// TIA Portal project "SMSS-ENLAB-01-003-1508-012-PLC-B_V13_SP1_1_V17" (V17) (continued)
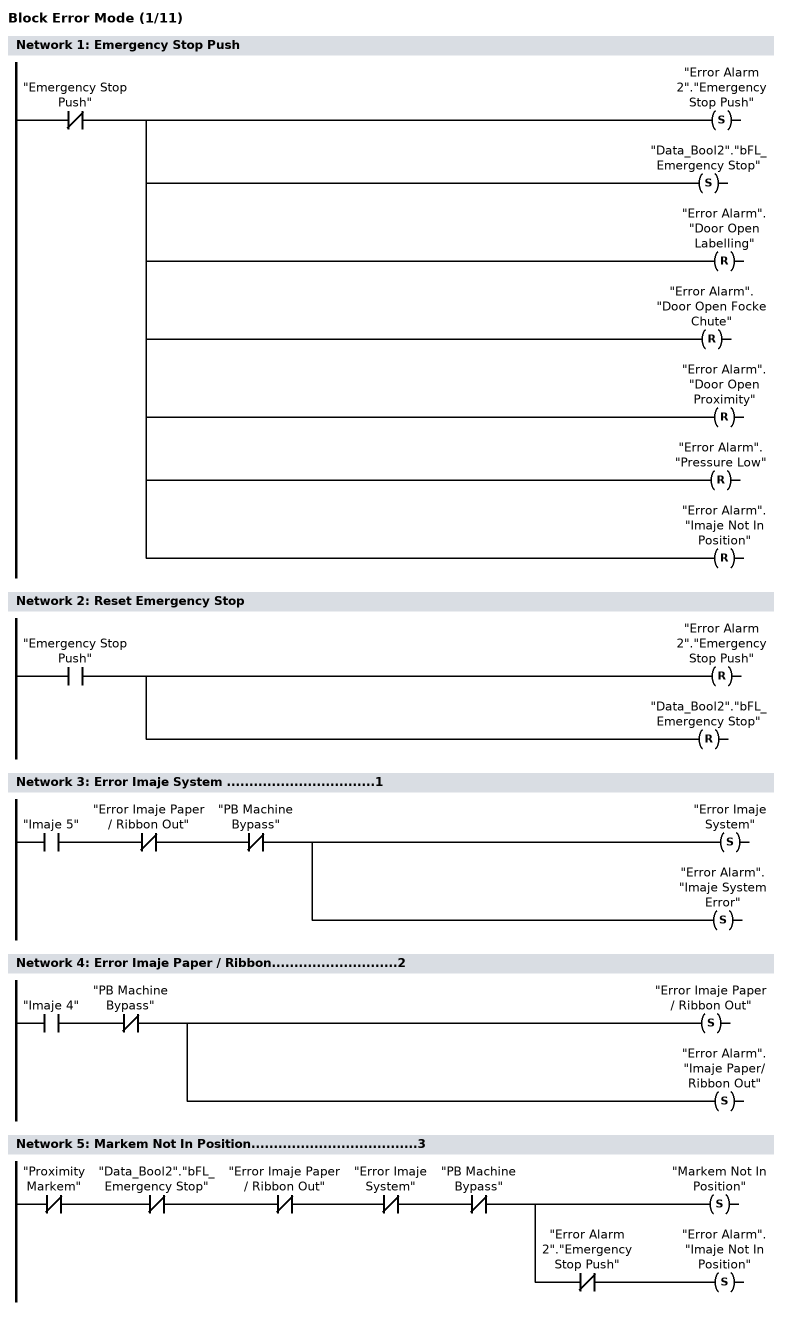
   RUNG wire#powerrail
      I_Contact( "Emergency Stop Push" )
      wire#w1
      S_Coil( "Error Alarm 2"."Emergency Stop Push" )
   END_RUNG
   RUNG wire#w1
      S_Coil( "Data_Bool2"."bFL_Emergency Stop" )
   END_RUNG
   RUNG wire#w1
      R_Coil( "Error Alarm"."Door Open Labelling" )
   END_RUNG
   RUNG wire#w1
      R_Coil( "Error Alarm"."Door Open Focke Chute" )
   END_RUNG
   RUNG wire#w1
      R_Coil( "Error Alarm"."Door Open Proximity" )
   END_RUNG
   RUNG wire#w1
      R_Coil( "Error Alarm"."Pressure Low" )
   END_RUNG
   RUNG wire#w1
      R_Coil( "Error Alarm"."Imaje Not In Position" )
   END_RUNG
   // the same network as SCL:
   IF NOT "Emergency Stop Push" THEN
       "Error Alarm 2"."Emergency Stop Push" := TRUE;
       "Data_Bool2"."bFL_Emergency Stop" := TRUE;
       "Error Alarm"."Door Open Labelling" := FALSE;
       "Error Alarm"."Door Open Focke Chute" := FALSE;
       "Error Alarm"."Door Open Proximity" := FALSE;
       "Error Alarm"."Pressure Low" := FALSE;
       "Error Alarm"."Imaje Not In Position" := FALSE;
   END_IF;
END_REGION

REGION Network 2: Reset Emergency Stop
   RUNG wire#powerrail
      Contact( "Emergency Stop Push" )
      wire#w1
      R_Coil( "Error Alarm 2"."Emergency Stop Push" )
   END_RUNG
   RUNG wire#w1
      R_Coil( "Data_Bool2"."bFL_Emergency Stop" )
   END_RUNG
   // the same network as SCL:
   IF "Emergency Stop Push" THEN
       "Error Alarm 2"."Emergency Stop Push" := FALSE;
       "Data_Bool2"."bFL_Emergency Stop" := FALSE;
   END_IF;
END_REGION

REGION Network 3: Error Imaje System .................................1
   RUNG wire#powerrail
      Contact( "Imaje 5" )
      I_Contact( "Error Imaje Paper / Ribbon Out" )
      I_Contact( "PB Machine Bypass" )
      wire#w1
      S_Coil( "Error Imaje System" )
   END_RUNG
   RUNG wire#w1
      S_Coil( "Error Alarm"."Imaje System Error" )
   END_RUNG
   // the same network as SCL:
   IF "Imaje 5" AND NOT "Error Imaje Paper / Ribbon Out" AND NOT "PB Machine Bypass" THEN
       "Error Imaje System" := TRUE;
       "Error Alarm"."Imaje System Error" := TRUE;
   END_IF;
END_REGION

REGION Network 4: Error Imaje Paper / Ribbon............................2
   RUNG wire#powerrail
      Contact( "Imaje 4" )
      I_Contact( "PB Machine Bypass" )
      wire#w1
      S_Coil( "Error Imaje Paper / Ribbon Out" )
   END_RUNG
   RUNG wire#w1
      S_Coil( "Error Alarm"."Imaje Paper/Ribbon Out" )
   END_RUNG
   // the same network as SCL:
   IF "Imaje 4" AND NOT "PB Machine Bypass" THEN
       "Error Imaje Paper / Ribbon Out" := TRUE;
       "Error Alarm"."Imaje Paper/Ribbon Out" := TRUE;
   END_IF;
END_REGION

REGION Network 5: Markem Not In Position.....................................3
   RUNG wire#powerrail
      I_Contact( "Proximity Markem" )
      I_Contact( "Data_Bool2"."bFL_Emergency Stop" )
      I_Contact( "Error Imaje Paper / Ribbon Out" )
      I_Contact( "Error Imaje System" )
      I_Contact( "PB Machine Bypass" )
      wire#w1
      S_Coil( "Markem Not In Position" )
   END_RUNG
   RUNG wire#w1
      I_Contact( "Error Alarm 2"."Emergency Stop Push" )
      S_Coil( "Error Alarm"."Imaje Not In Position" )
   END_RUNG
   // the same network as SCL:
   #_w1 := NOT "Proximity Markem" AND NOT "Data_Bool2"."bFL_Emergency Stop" AND NOT "Error Imaje Paper / Ribbon Out" AND NOT "Error Imaje System" AND NOT "PB Machine Bypass";
   IF #_w1 THEN "Markem Not In Position" := TRUE; END_IF;
   IF #_w1 AND NOT "Error Alarm 2"."Emergency Stop Push" THEN
       "Error Alarm"."Imaje Not In Position" := TRUE;
   END_IF;
END_REGION

REGION Network 6: Groub Error Imaje Jika baypass mesin Off
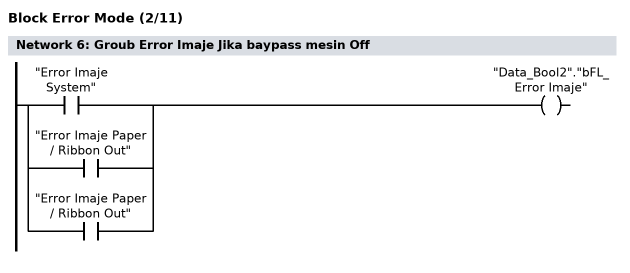
   RUNG wire#powerrail
      Contact( "Error Imaje System" )
      wire#w1
      Coil( "Data_Bool2"."bFL_Error Imaje" )
   END_RUNG
   RUNG wire#powerrail
      Contact( "Error Imaje Paper / Ribbon Out" )
   END_RUNG wire#w1
   RUNG wire#powerrail
      Contact( "Error Imaje Paper / Ribbon Out" )
   END_RUNG wire#w1
   // the same network as SCL:
   "Data_Bool2"."bFL_Error Imaje" := "Error Imaje System" OR "Error Imaje Paper / Ribbon Out" OR "Error Imaje Paper / Ribbon Out";
END_REGION

REGION Network 7: Error Imaje Reset Other Error
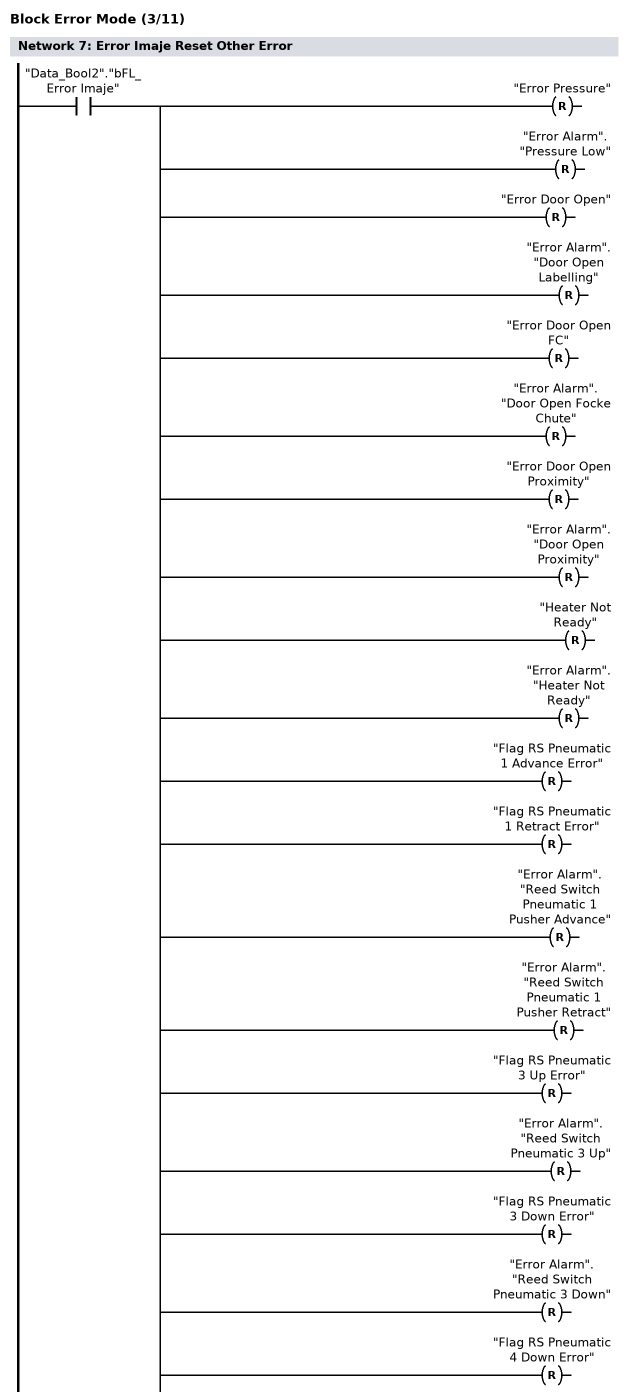
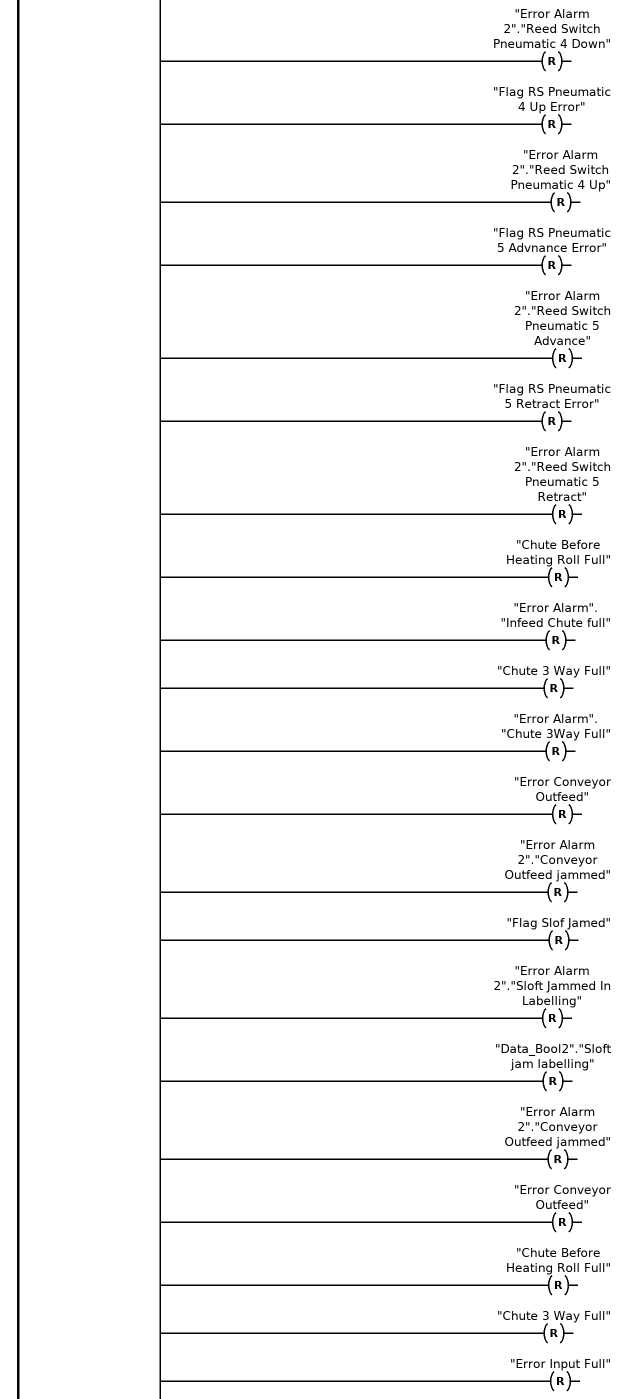
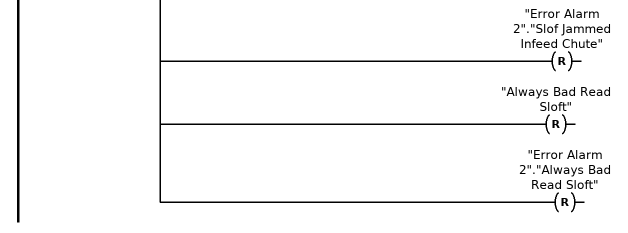
   RUNG wire#powerrail
      Contact( "Data_Bool2"."bFL_Error Imaje" )
      wire#w1
      R_Coil( "Error Pressure" )
   END_RUNG
   RUNG wire#w1
      R_Coil( "Error Alarm"."Pressure Low" )
   END_RUNG
   RUNG wire#w1
      R_Coil( "Error Door Open" )
   END_RUNG
   RUNG wire#w1
      R_Coil( "Error Alarm"."Door Open Labelling" )
   END_RUNG
   RUNG wire#w1
      R_Coil( "Error Door Open FC" )
   END_RUNG
   RUNG wire#w1
      R_Coil( "Error Alarm"."Door Open Focke Chute" )
   END_RUNG
   RUNG wire#w1
      R_Coil( "Error Door Open Proximity" )
   END_RUNG
   RUNG wire#w1
      R_Coil( "Error Alarm"."Door Open Proximity" )
   END_RUNG
   RUNG wire#w1
      R_Coil( "Heater Not Ready" )
   END_RUNG
   RUNG wire#w1
      R_Coil( "Error Alarm"."Heater Not Ready" )
   END_RUNG
   RUNG wire#w1
      R_Coil( "Flag RS Pneumatic 1 Advance Error" )
   END_RUNG
   RUNG wire#w1
      R_Coil( "Flag RS Pneumatic 1 Retract Error" )
   END_RUNG
   RUNG wire#w1
      R_Coil( "Error Alarm"."Reed Switch Pneumatic 1 Pusher Advance" )
   END_RUNG
   RUNG wire#w1
      R_Coil( "Error Alarm"."Reed Switch Pneumatic 1 Pusher Retract" )
   END_RUNG
   RUNG wire#w1
      R_Coil( "Flag RS Pneumatic 3 Up Error" )
   END_RUNG
   RUNG wire#w1
      R_Coil( "Error Alarm"."Reed Switch Pneumatic 3 Up" )
   END_RUNG
   RUNG wire#w1
      R_Coil( "Flag RS Pneumatic 3 Down Error" )
   END_RUNG
   RUNG wire#w1
      R_Coil( "Error Alarm"."Reed Switch Pneumatic 3 Down" )
   END_RUNG
   RUNG wire#w1
      R_Coil( "Flag RS Pneumatic 4 Down Error" )
   END_RUNG
   RUNG wire#w1
      R_Coil( "Error Alarm 2"."Reed Switch Pneumatic 4 Down" )
   END_RUNG
   RUNG wire#w1
      R_Coil( "Flag RS Pneumatic 4 Up Error" )
   END_RUNG
   RUNG wire#w1
      R_Coil( "Error Alarm 2"."Reed Switch Pneumatic 4 Up" )
   END_RUNG
   RUNG wire#w1
      R_Coil( "Flag RS Pneumatic 5 Advnance Error" )
   END_RUNG
   RUNG wire#w1
      R_Coil( "Error Alarm 2"."Reed Switch Pneumatic 5 Advance" )
   END_RUNG
   RUNG wire#w1
      R_Coil( "Flag RS Pneumatic 5 Retract Error" )
   END_RUNG
   RUNG wire#w1
      R_Coil( "Error Alarm 2"."Reed Switch Pneumatic 5 Retract" )
   END_RUNG
   RUNG wire#w1
      R_Coil( "Chute Before Heating Roll Full" )
   END_RUNG
   RUNG wire#w1
      R_Coil( "Error Alarm"."Infeed Chute full" )
   END_RUNG
   RUNG wire#w1
      R_Coil( "Chute 3 Way Full" )
   END_RUNG
   RUNG wire#w1
      R_Coil( "Error Alarm"."Chute 3Way Full" )
   END_RUNG
   RUNG wire#w1
      R_Coil( "Error Conveyor Outfeed" )
   END_RUNG
   RUNG wire#w1
      R_Coil( "Error Alarm 2"."Conveyor Outfeed jammed" )
   END_RUNG
   RUNG wire#w1
      R_Coil( "Flag Slof Jamed" )
   END_RUNG
   RUNG wire#w1
      R_Coil( "Error Alarm 2"."Sloft Jammed In Labelling" )
   END_RUNG
   RUNG wire#w1
      R_Coil( "Data_Bool2"."Sloft jam labelling" )
   END_RUNG
   RUNG wire#w1
      R_Coil( "Error Alarm 2"."Conveyor Outfeed jammed" )
   END_RUNG
   RUNG wire#w1
      R_Coil( "Error Conveyor Outfeed" )
   END_RUNG
   RUNG wire#w1
      R_Coil( "Chute Before Heating Roll Full" )
   END_RUNG
   RUNG wire#w1
      R_Coil( "Chute 3 Way Full" )
   END_RUNG
   RUNG wire#w1
      R_Coil( "Error Input Full" )
   END_RUNG
   RUNG wire#w1
      R_Coil( "Error Alarm 2"."Slof Jammed Infeed Chute" )
   END_RUNG
   RUNG wire#w1
      R_Coil( "Always Bad Read Sloft" )
   END_RUNG
   RUNG wire#w1
      R_Coil( "Error Alarm 2"."Always Bad Read Sloft" )
   END_RUNG
   // the same network as SCL:
   IF "Data_Bool2"."bFL_Error Imaje" THEN
       "Error Pressure" := FALSE;
       "Error Alarm"."Pressure Low" := FALSE;
       "Error Door Open" := FALSE;
       "Error Alarm"."Door Open Labelling" := FALSE;
       "Error Door Open FC" := FALSE;
       "Error Alarm"."Door Open Focke Chute" := FALSE;
       "Error Door Open Proximity" := FALSE;
       "Error Alarm"."Door Open Proximity" := FALSE;
       "Heater Not Ready" := FALSE;
       "Error Alarm"."Heater Not Ready" := FALSE;
       "Flag RS Pneumatic 1 Advance Error" := FALSE;
       "Flag RS Pneumatic 1 Retract Error" := FALSE;
       "Error Alarm"."Reed Switch Pneumatic 1 Pusher Advance" := FALSE;
       "Error Alarm"."Reed Switch Pneumatic 1 Pusher Retract" := FALSE;
       "Flag RS Pneumatic 3 Up Error" := FALSE;
       "Error Alarm"."Reed Switch Pneumatic 3 Up" := FALSE;
       "Flag RS Pneumatic 3 Down Error" := FALSE;
       "Error Alarm"."Reed Switch Pneumatic 3 Down" := FALSE;
       "Flag RS Pneumatic 4 Down Error" := FALSE;
       "Error Alarm 2"."Reed Switch Pneumatic 4 Down" := FALSE;
       "Flag RS Pneumatic 4 Up Error" := FALSE;
       "Error Alarm 2"."Reed Switch Pneumatic 4 Up" := FALSE;
       "Flag RS Pneumatic 5 Advnance Error" := FALSE;
       "Error Alarm 2"."Reed Switch Pneumatic 5 Advance" := FALSE;
       "Flag RS Pneumatic 5 Retract Error" := FALSE;
       "Error Alarm 2"."Reed Switch Pneumatic 5 Retract" := FALSE;
       "Chute Before Heating Roll Full" := FALSE;
       "Error Alarm"."Infeed Chute full" := FALSE;
       "Chute 3 Way Full" := FALSE;
       "Error Alarm"."Chute 3Way Full" := FALSE;
       "Error Conveyor Outfeed" := FALSE;
       "Error Alarm 2"."Conveyor Outfeed jammed" := FALSE;
       "Flag Slof Jamed" := FALSE;
       "Error Alarm 2"."Sloft Jammed In Labelling" := FALSE;
       "Data_Bool2"."Sloft jam labelling" := FALSE;
       "Error Alarm 2"."Conveyor Outfeed jammed" := FALSE;
       "Error Conveyor Outfeed" := FALSE;
       "Chute Before Heating Roll Full" := FALSE;
       "Chute 3 Way Full" := FALSE;
       "Error Input Full" := FALSE;
       "Error Alarm 2"."Slof Jammed Infeed Chute" := FALSE;
       "Always Bad Read Sloft" := FALSE;
       "Error Alarm 2"."Always Bad Read Sloft" := FALSE;
   END_IF;
END_REGION

REGION Network 8: Other Error Imaje Reset Error Imaje
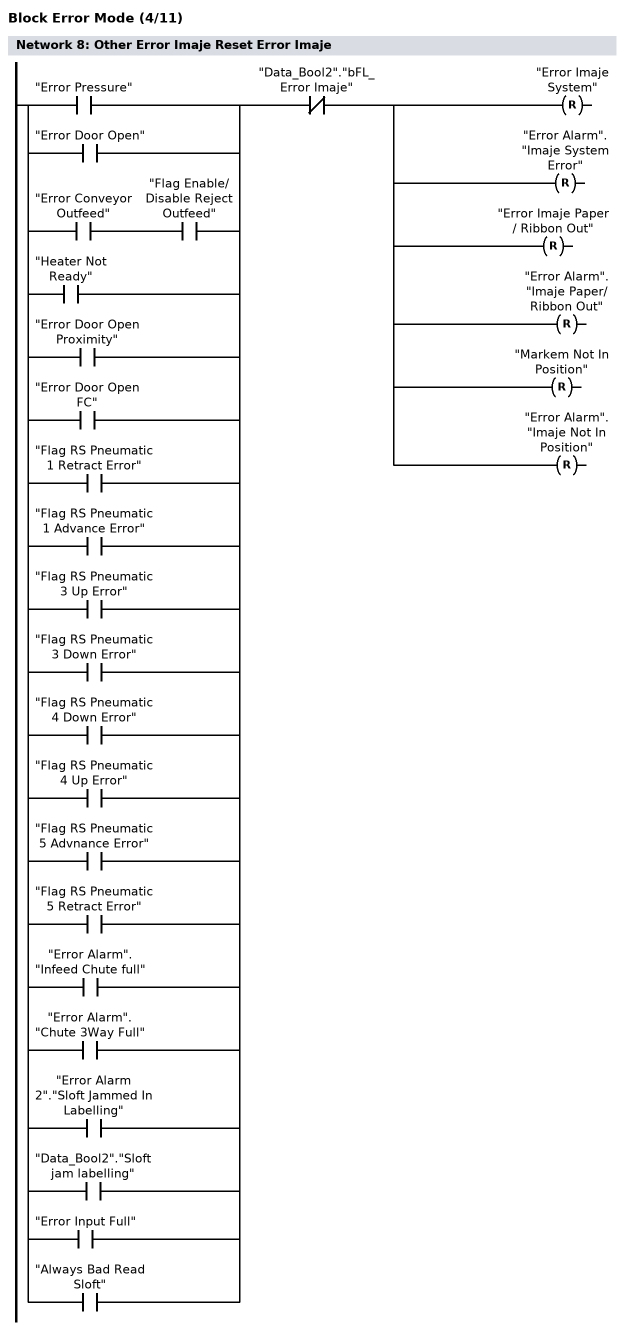
   RUNG wire#powerrail
      Contact( "Error Pressure" )
      wire#w1
      I_Contact( "Data_Bool2"."bFL_Error Imaje" )
      wire#w2
      R_Coil( "Error Imaje System" )
   END_RUNG
   RUNG wire#powerrail
      Contact( "Error Door Open" )
   END_RUNG wire#w1
   RUNG wire#powerrail
      Contact( "Error Conveyor Outfeed" )
      Contact( "Flag Enable/Disable Reject Outfeed" )
   END_RUNG wire#w1
   RUNG wire#powerrail
      Contact( "Heater Not Ready" )
   END_RUNG wire#w1
   RUNG wire#powerrail
      Contact( "Error Door Open Proximity" )
   END_RUNG wire#w1
   RUNG wire#powerrail
      Contact( "Error Door Open FC" )
   END_RUNG wire#w1
   RUNG wire#powerrail
      Contact( "Flag RS Pneumatic 1 Retract Error" )
   END_RUNG wire#w1
   RUNG wire#powerrail
      Contact( "Flag RS Pneumatic 1 Advance Error" )
   END_RUNG wire#w1
   RUNG wire#powerrail
      Contact( "Flag RS Pneumatic 3 Up Error" )
   END_RUNG wire#w1
   RUNG wire#powerrail
      Contact( "Flag RS Pneumatic 3 Down Error" )
   END_RUNG wire#w1
   RUNG wire#powerrail
      Contact( "Flag RS Pneumatic 4 Down Error" )
   END_RUNG wire#w1
   RUNG wire#powerrail
      Contact( "Flag RS Pneumatic 4 Up Error" )
   END_RUNG wire#w1
   RUNG wire#powerrail
      Contact( "Flag RS Pneumatic 5 Advnance Error" )
   END_RUNG wire#w1
   RUNG wire#powerrail
      Contact( "Flag RS Pneumatic 5 Retract Error" )
   END_RUNG wire#w1
   RUNG wire#powerrail
      Contact( "Error Alarm"."Infeed Chute full" )
   END_RUNG wire#w1
   RUNG wire#powerrail
      Contact( "Error Alarm"."Chute 3Way Full" )
   END_RUNG wire#w1
   RUNG wire#powerrail
      Contact( "Error Alarm 2"."Sloft Jammed In Labelling" )
   END_RUNG wire#w1
   RUNG wire#powerrail
      Contact( "Data_Bool2"."Sloft jam labelling" )
   END_RUNG wire#w1
   RUNG wire#powerrail
      Contact( "Error Input Full" )
   END_RUNG wire#w1
   RUNG wire#powerrail
      Contact( "Always Bad Read Sloft" )
   END_RUNG wire#w1
   RUNG wire#w2
      R_Coil( "Error Alarm"."Imaje System Error" )
   END_RUNG
   RUNG wire#w2
      R_Coil( "Error Imaje Paper / Ribbon Out" )
   END_RUNG
   RUNG wire#w2
      R_Coil( "Error Alarm"."Imaje Paper/Ribbon Out" )
   END_RUNG
   RUNG wire#w2
      R_Coil( "Markem Not In Position" )
   END_RUNG
   RUNG wire#w2
      R_Coil( "Error Alarm"."Imaje Not In Position" )
   END_RUNG
   // the same network as SCL:
   IF ("Error Pressure" OR "Error Door Open" OR ("Error Conveyor Outfeed" AND "Flag Enable/Disable Reject Outfeed") OR "Heater Not Ready" OR "Error Door Open Proximity" OR "Error Door Open FC" OR "Flag RS Pneumatic 1 Retract Error" OR "Flag RS Pneumatic 1 Advance Error" OR "Flag RS Pneumatic 3 Up Error" OR "Flag RS Pneumatic 3 Down Error" OR "Flag RS Pneumatic 4 Down Error" OR "Flag RS Pneumatic 4 Up Error" OR "Flag RS Pneumatic 5 Advnance Error" OR "Flag RS Pneumatic 5 Retract Error" OR "Error Alarm"."Infeed Chute full" OR "Error Alarm"."Chute 3Way Full" OR "Error Alarm 2"."Sloft Jammed In Labelling" OR "Data_Bool2"."Sloft jam labelling" OR "Error Input Full" OR "Always Bad Read Sloft") AND NOT "Data_Bool2"."bFL_Error Imaje" THEN
       "Error Imaje System" := FALSE;
       "Error Alarm"."Imaje System Error" := FALSE;
       "Error Imaje Paper / Ribbon Out" := FALSE;
       "Error Alarm"."Imaje Paper/Ribbon Out" := FALSE;
       "Markem Not In Position" := FALSE;
       "Error Alarm"."Imaje Not In Position" := FALSE;
   END_IF;
END_REGION

REGION Network 9: Set Bad Read Berturut-rurut -----------> mesin Error ..................................4
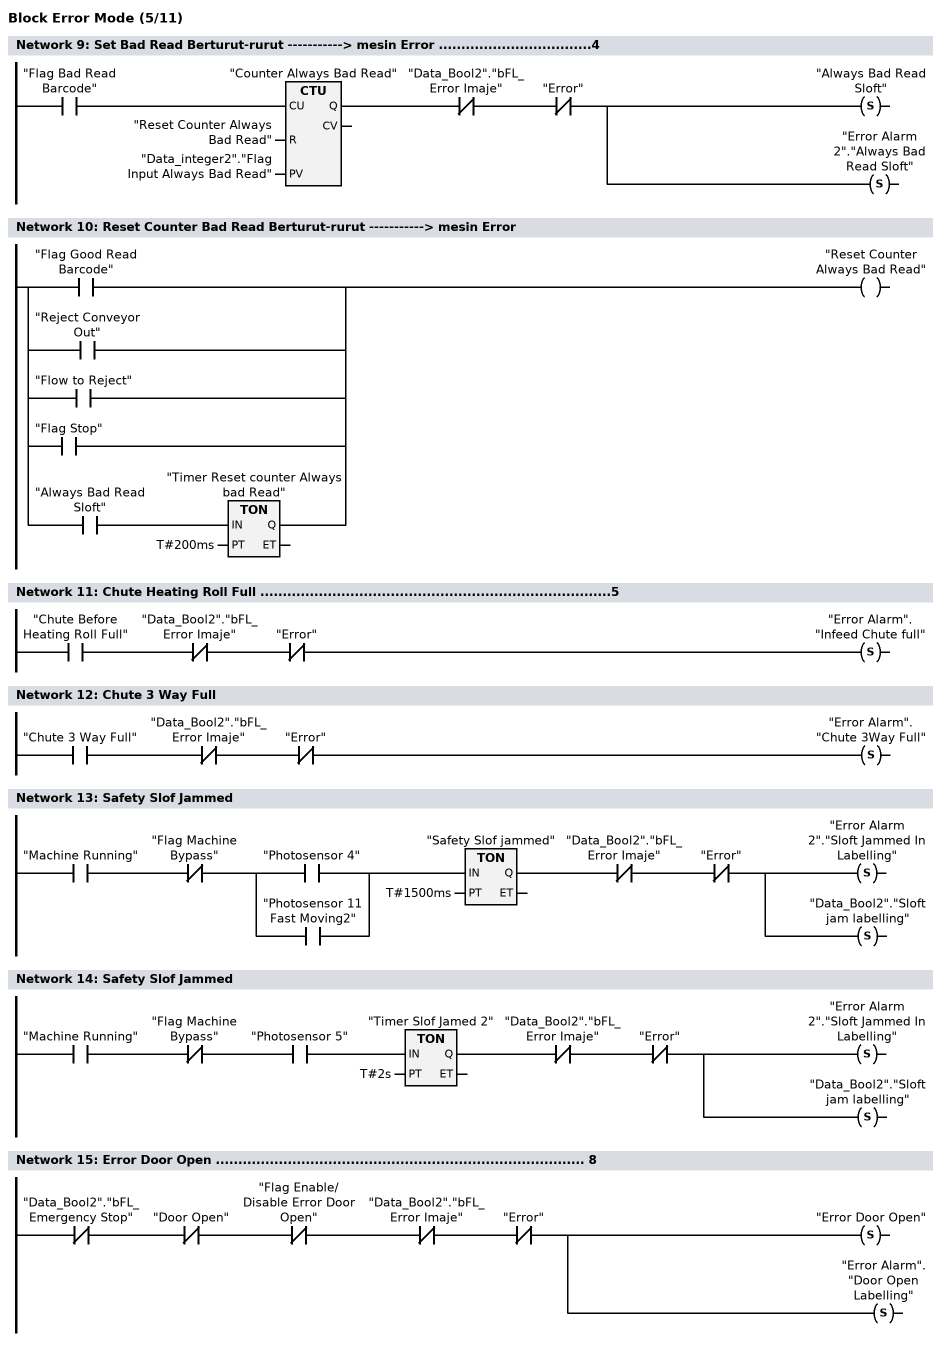
   "Counter Always Bad Read".CTU(CU := "Flag Bad Read Barcode",
                           R := "Reset Counter Always Bad Read",
                           PV := "Data_integer2"."Flag Input Always Bad Read");
   IF "Counter Always Bad Read".Q AND NOT "Data_Bool2"."bFL_Error Imaje" AND NOT "Error" THEN
       "Always Bad Read Sloft" := TRUE;
       "Error Alarm 2"."Always Bad Read Sloft" := TRUE;
   END_IF;
END_REGION

REGION Network 10: Reset Counter Bad Read Berturut-rurut -----------> mesin Error
   "Timer Reset counter Always bad Read".TON(IN := "Always Bad Read Sloft", PT := T#200ms);
   "Reset Counter Always Bad Read" := "Flag Good Read Barcode" OR "Reject Conveyor Out" OR "Flow to Reject" OR "Flag Stop" OR "Timer Reset counter Always bad Read".Q;
END_REGION

REGION Network 11: Chute Heating Roll Full ..............................................................................5
   RUNG wire#powerrail
      Contact( "Chute Before Heating Roll Full" )
      I_Contact( "Data_Bool2"."bFL_Error Imaje" )
      I_Contact( "Error" )
      S_Coil( "Error Alarm"."Infeed Chute full" )
   END_RUNG
   // the same network as SCL:
   IF "Chute Before Heating Roll Full" AND NOT "Data_Bool2"."bFL_Error Imaje" AND NOT "Error" THEN
       "Error Alarm"."Infeed Chute full" := TRUE;
   END_IF;
END_REGION

REGION Network 12: Chute 3 Way Full
   RUNG wire#powerrail
      Contact( "Chute 3 Way Full" )
      I_Contact( "Data_Bool2"."bFL_Error Imaje" )
      I_Contact( "Error" )
      S_Coil( "Error Alarm"."Chute 3Way Full" )
   END_RUNG
   // the same network as SCL:
   IF "Chute 3 Way Full" AND NOT "Data_Bool2"."bFL_Error Imaje" AND NOT "Error" THEN
       "Error Alarm"."Chute 3Way Full" := TRUE;
   END_IF;
END_REGION

REGION Network 13: Safety Slof Jammed
   "Safety Slof jammed".TON(IN := "Machine Running" AND NOT "Flag Machine Bypass" AND ("Photosensor 4" OR "Photosensor 11 Fast Moving2"),
                           PT := T#1500ms);
   IF "Safety Slof jammed".Q AND NOT "Data_Bool2"."bFL_Error Imaje" AND NOT "Error" THEN
       "Error Alarm 2"."Sloft Jammed In Labelling" := TRUE;
       "Data_Bool2"."Sloft jam labelling" := TRUE;
   END_IF;
END_REGION

REGION Network 14: Safety Slof Jammed
   "Timer Slof Jamed 2".TON(IN := "Machine Running" AND NOT "Flag Machine Bypass" AND "Photosensor 5",
                           PT := T#2s);
   IF "Timer Slof Jamed 2".Q AND NOT "Data_Bool2"."bFL_Error Imaje" AND NOT "Error" THEN
       "Error Alarm 2"."Sloft Jammed In Labelling" := TRUE;
       "Data_Bool2"."Sloft jam labelling" := TRUE;
   END_IF;
END_REGION

REGION Network 15: Error Door Open .................................................................................. 8
   RUNG wire#powerrail
      I_Contact( "Data_Bool2"."bFL_Emergency Stop" )
      I_Contact( "Door Open" )
      I_Contact( "Flag Enable/Disable Error Door Open" )
      I_Contact( "Data_Bool2"."bFL_Error Imaje" )
      I_Contact( "Error" )
      wire#w1
      S_Coil( "Error Door Open" )
   END_RUNG
   RUNG wire#w1
      S_Coil( "Error Alarm"."Door Open Labelling" )
   END_RUNG
   // the same network as SCL:
   IF NOT "Data_Bool2"."bFL_Emergency Stop" AND NOT "Door Open" AND NOT "Flag Enable/Disable Error Door Open" AND NOT "Data_Bool2"."bFL_Error Imaje" AND NOT "Error" THEN
       "Error Door Open" := TRUE;
       "Error Alarm"."Door Open Labelling" := TRUE;
   END_IF;
END_REGION

REGION Network 16: Error Door Open FC
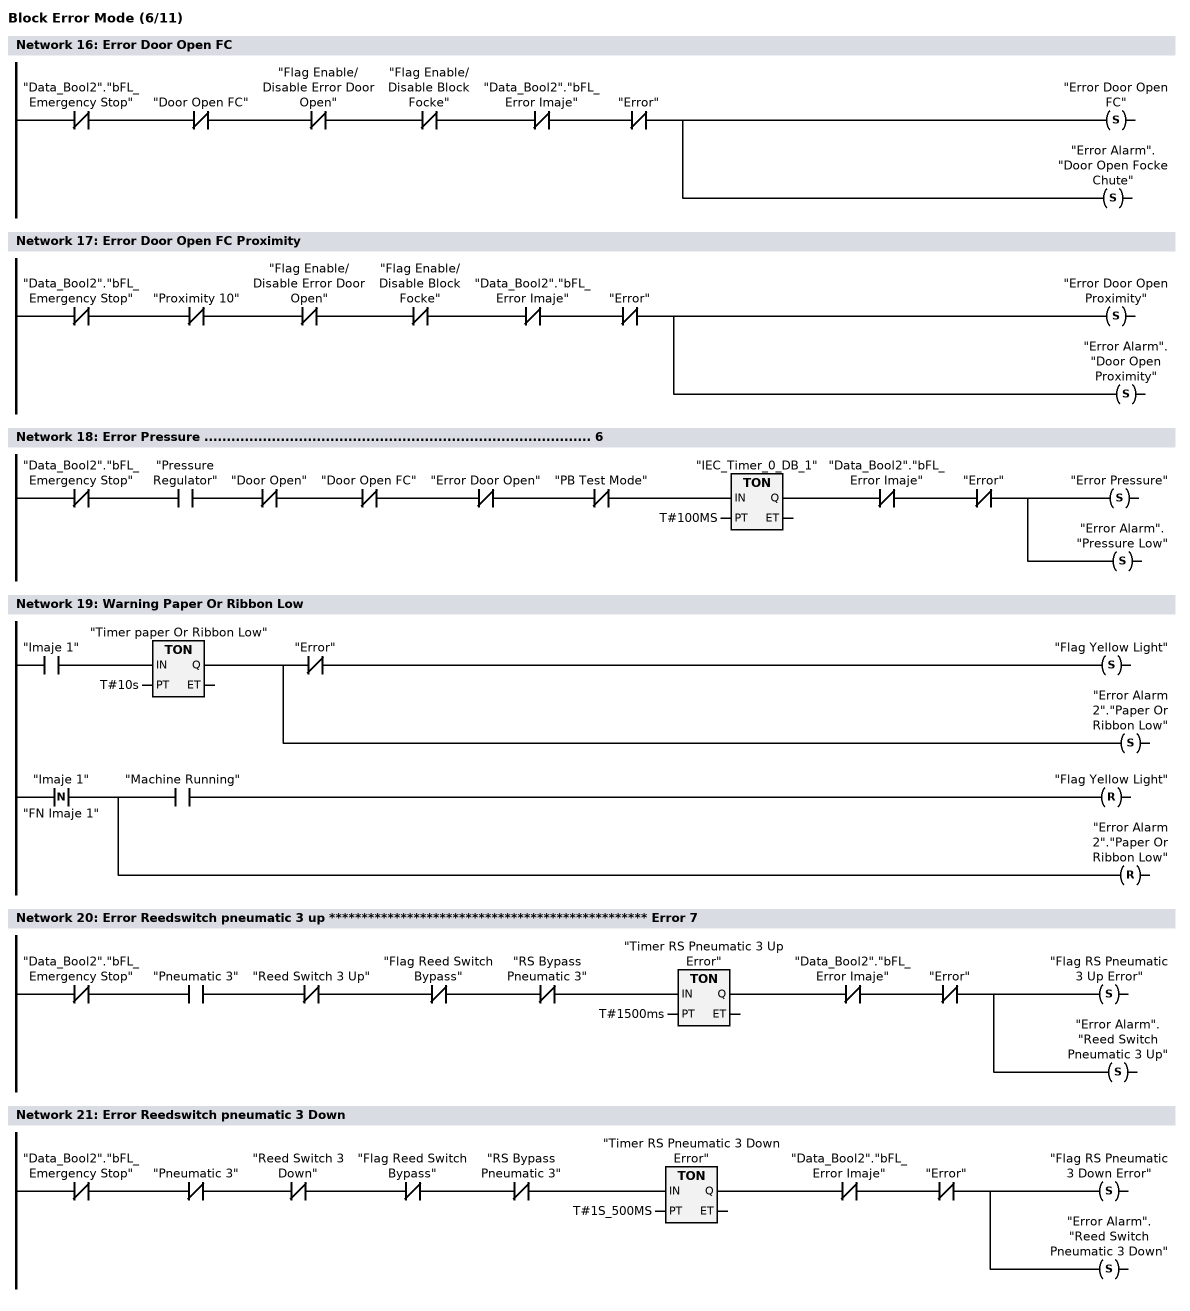
   RUNG wire#powerrail
      I_Contact( "Data_Bool2"."bFL_Emergency Stop" )
      I_Contact( "Door Open FC" )
      I_Contact( "Flag Enable/Disable Error Door Open" )
      I_Contact( "Flag Enable/Disable Block Focke" )
      I_Contact( "Data_Bool2"."bFL_Error Imaje" )
      I_Contact( "Error" )
      wire#w1
      S_Coil( "Error Door Open FC" )
   END_RUNG
   RUNG wire#w1
      S_Coil( "Error Alarm"."Door Open Focke Chute" )
   END_RUNG
   // the same network as SCL:
   IF NOT "Data_Bool2"."bFL_Emergency Stop" AND NOT "Door Open FC" AND NOT "Flag Enable/Disable Error Door Open" AND NOT "Flag Enable/Disable Block Focke" AND NOT "Data_Bool2"."bFL_Error Imaje" AND NOT "Error" THEN
       "Error Door Open FC" := TRUE;
       "Error Alarm"."Door Open Focke Chute" := TRUE;
   END_IF;
END_REGION

REGION Network 17: Error Door Open FC Proximity
   RUNG wire#powerrail
      I_Contact( "Data_Bool2"."bFL_Emergency Stop" )
      I_Contact( "Proximity 10" )
      I_Contact( "Flag Enable/Disable Error Door Open" )
      I_Contact( "Flag Enable/Disable Block Focke" )
      I_Contact( "Data_Bool2"."bFL_Error Imaje" )
      I_Contact( "Error" )
      wire#w1
      S_Coil( "Error Door Open Proximity" )
   END_RUNG
   RUNG wire#w1
      S_Coil( "Error Alarm"."Door Open Proximity" )
   END_RUNG
   // the same network as SCL:
   IF NOT "Data_Bool2"."bFL_Emergency Stop" AND NOT "Proximity 10" AND NOT "Flag Enable/Disable Error Door Open" AND NOT "Flag Enable/Disable Block Focke" AND NOT "Data_Bool2"."bFL_Error Imaje" AND NOT "Error" THEN
       "Error Door Open Proximity" := TRUE;
       "Error Alarm"."Door Open Proximity" := TRUE;
   END_IF;
END_REGION

REGION Network 18: Error Pressure ...................................................................................... 6
   "IEC_Timer_0_DB_1".TON(IN := NOT "Data_Bool2"."bFL_Emergency Stop" AND "Pressure Regulator" AND NOT "Door Open" AND NOT "Door Open FC" AND NOT "Error Door Open" AND NOT "PB Test Mode",
                          PT := T#100MS);
   IF "IEC_Timer_0_DB_1".Q AND NOT "Data_Bool2"."bFL_Error Imaje" AND NOT "Error" THEN
       "Error Pressure" := TRUE;
       "Error Alarm"."Pressure Low" := TRUE;
   END_IF;
END_REGION

REGION Network 19: Warning Paper Or Ribbon Low
   "Timer paper Or Ribbon Low".TON(IN := "Imaje 1", PT := T#10s);
   IF "Timer paper Or Ribbon Low".Q AND NOT "Error" THEN "Flag Yellow Light" := TRUE; END_IF;
   IF "Timer paper Or Ribbon Low".Q THEN "Error Alarm 2"."Paper Or Ribbon Low" := TRUE; END_IF;
   #_w1 := NOT "Imaje 1" AND "FN Imaje 1";   // falling edge of "Imaje 1"
   "FN Imaje 1" := "Imaje 1";
   IF #_w1 AND "Machine Running" THEN "Flag Yellow Light" := FALSE; END_IF;
   IF #_w1 THEN "Error Alarm 2"."Paper Or Ribbon Low" := FALSE; END_IF;
END_REGION

REGION Network 20: Error Reedswitch pneumatic 3 up ************************************************* Error 7
   "Timer RS Pneumatic 3 Up Error".TON(IN := NOT "Data_Bool2"."bFL_Emergency Stop" AND "Pneumatic 3" AND NOT "Reed Switch 3 Up" AND NOT "Flag Reed Switch Bypass" AND NOT "RS Bypass Pneumatic 3",
                           PT := T#1500ms);
   IF "Timer RS Pneumatic 3 Up Error".Q AND NOT "Data_Bool2"."bFL_Error Imaje" AND NOT "Error" THEN
       "Flag RS Pneumatic 3 Up Error" := TRUE;
       "Error Alarm"."Reed Switch Pneumatic 3 Up" := TRUE;
   END_IF;
END_REGION

REGION Network 21: Error Reedswitch pneumatic 3 Down
   "Timer RS Pneumatic 3 Down Error".TON(IN := NOT "Data_Bool2"."bFL_Emergency Stop" AND NOT "Pneumatic 3" AND NOT "Reed Switch 3 Down" AND NOT "Flag Reed Switch Bypass" AND NOT "RS Bypass Pneumatic 3",
                           PT := T#1S_500MS);
   IF "Timer RS Pneumatic 3 Down Error".Q AND NOT "Data_Bool2"."bFL_Error Imaje" AND NOT "Error" THEN
       "Flag RS Pneumatic 3 Down Error" := TRUE;
       "Error Alarm"."Reed Switch Pneumatic 3 Down" := TRUE;
   END_IF;
END_REGION

REGION Network 22: Error Reedswitch pneumatic 4 Down
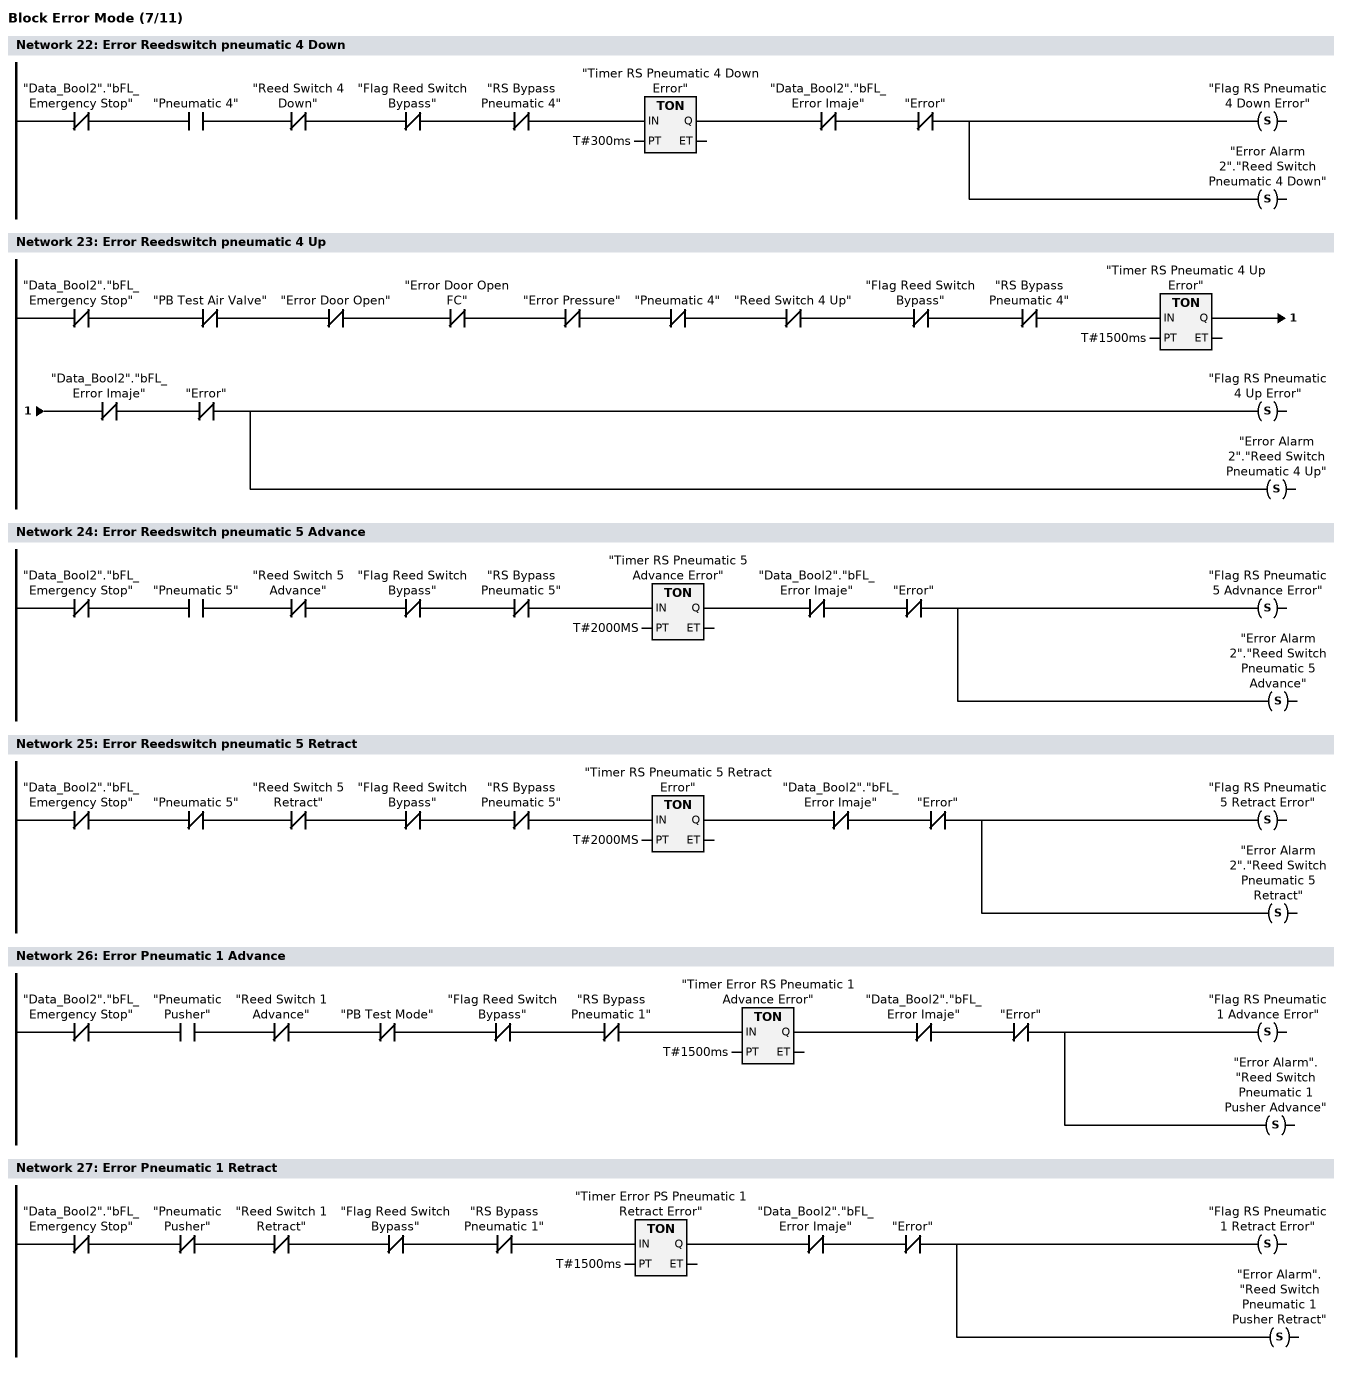
   "Timer RS Pneumatic 4 Down Error".TON(IN := NOT "Data_Bool2"."bFL_Emergency Stop" AND "Pneumatic 4" AND NOT "Reed Switch 4 Down" AND NOT "Flag Reed Switch Bypass" AND NOT "RS Bypass Pneumatic 4",
                           PT := T#300ms);
   IF "Timer RS Pneumatic 4 Down Error".Q AND NOT "Data_Bool2"."bFL_Error Imaje" AND NOT "Error" THEN
       "Flag RS Pneumatic 4 Down Error" := TRUE;
       "Error Alarm 2"."Reed Switch Pneumatic 4 Down" := TRUE;
   END_IF;
END_REGION

REGION Network 23: Error Reedswitch pneumatic 4 Up
   "Timer RS Pneumatic 4 Up Error".TON(IN := NOT "Data_Bool2"."bFL_Emergency Stop" AND NOT "PB Test Air Valve" AND NOT "Error Door Open" AND NOT "Error Door Open FC" AND NOT "Error Pressure" AND NOT "Pneumatic 4" AND NOT "Reed Switch 4 Up" AND NOT "Flag Reed Switch Bypass" AND NOT "RS Bypass Pneumatic 4",
                           PT := T#1500ms);
   IF "Timer RS Pneumatic 4 Up Error".Q AND NOT "Data_Bool2"."bFL_Error Imaje" AND NOT "Error" THEN
       "Flag RS Pneumatic 4 Up Error" := TRUE;
       "Error Alarm 2"."Reed Switch Pneumatic 4 Up" := TRUE;
   END_IF;
END_REGION

REGION Network 24: Error Reedswitch pneumatic 5 Advance
   "Timer RS Pneumatic 5 Advance Error".TON(IN := NOT "Data_Bool2"."bFL_Emergency Stop" AND "Pneumatic 5" AND NOT "Reed Switch 5 Advance" AND NOT "Flag Reed Switch Bypass" AND NOT "RS Bypass Pneumatic 5",
                           PT := T#2000MS);
   IF "Timer RS Pneumatic 5 Advance Error".Q AND NOT "Data_Bool2"."bFL_Error Imaje" AND NOT "Error" THEN
       "Flag RS Pneumatic 5 Advnance Error" := TRUE;
       "Error Alarm 2"."Reed Switch Pneumatic 5 Advance" := TRUE;
   END_IF;
END_REGION

REGION Network 25: Error Reedswitch pneumatic 5 Retract
   "Timer RS Pneumatic 5 Retract Error".TON(IN := NOT "Data_Bool2"."bFL_Emergency Stop" AND NOT "Pneumatic 5" AND NOT "Reed Switch 5 Retract" AND NOT "Flag Reed Switch Bypass" AND NOT "RS Bypass Pneumatic 5",
                           PT := T#2000MS);
   IF "Timer RS Pneumatic 5 Retract Error".Q AND NOT "Data_Bool2"."bFL_Error Imaje" AND NOT "Error" THEN
       "Flag RS Pneumatic 5 Retract Error" := TRUE;
       "Error Alarm 2"."Reed Switch Pneumatic 5 Retract" := TRUE;
   END_IF;
END_REGION

REGION Network 26: Error Pneumatic 1 Advance
   "Timer Error RS Pneumatic 1 Advance Error".TON(IN := NOT "Data_Bool2"."bFL_Emergency Stop" AND "Pneumatic Pusher" AND NOT "Reed Switch 1 Advance" AND NOT "PB Test Mode" AND NOT "Flag Reed Switch Bypass" AND NOT "RS Bypass Pneumatic 1",
                           PT := T#1500ms);
   IF "Timer Error RS Pneumatic 1 Advance Error".Q AND NOT "Data_Bool2"."bFL_Error Imaje" AND NOT "Error" THEN
       "Flag RS Pneumatic 1 Advance Error" := TRUE;
       "Error Alarm"."Reed Switch Pneumatic 1 Pusher Advance" := TRUE;
   END_IF;
END_REGION

REGION Network 27: Error Pneumatic 1 Retract
   "Timer Error PS Pneumatic 1 Retract Error".TON(IN := NOT "Data_Bool2"."bFL_Emergency Stop" AND NOT "Pneumatic Pusher" AND NOT "Reed Switch 1 Retract" AND NOT "Flag Reed Switch Bypass" AND NOT "RS Bypass Pneumatic 1",
                           PT := T#1500ms);
   IF "Timer Error PS Pneumatic 1 Retract Error".Q AND NOT "Data_Bool2"."bFL_Error Imaje" AND NOT "Error" THEN
       "Flag RS Pneumatic 1 Retract Error" := TRUE;
       "Error Alarm"."Reed Switch Pneumatic 1 Pusher Retract" := TRUE;
   END_IF;
END_REGION

REGION Network 28: All Error
   // Semua Error